// TIA Portal project "TNprojINZ" (V15.1) (continued)

       ELSIF ("OPC - z LabVIEW"."Poziom zbiornik 4" > ("OPC - do LabVIEW"."PRO poziom cieczy Z4" + 3)) THEN
           "OPC - do LabVIEW"."Zawór spustowy Z4" := 1;
           "Z4 globalne"."Czy Z4 pełny?" := 0;

       ELSIF ("OPC - z LabVIEW"."Poziom zbiornik 4" < ("OPC - do LabVIEW"."PRO poziom cieczy Z4" - 3)) THEN
           "OPC - do LabVIEW"."Zawór spustowy Z4" := 0;
           "Z4 globalne"."Czy Z4 pełny?" := 0;
       END_IF;
   //ELSE
       //"Z4 globalne"."Czy Z4 pełny?" := 0;
   END_IF;
END_FUNCTION_BLOCK

FUNCTION_BLOCK "SCL - Grzanie"   // FB9, SCL
{ S7_Optimized_Access := 'TRUE' }
VERSION : 0.1
BEGIN
   (*
   4 x - dla każdego zbiornika oddzielnie 
   if then               i Awaria = 0
       proces grzania
   else - koniec proc grz
       reset - "Z1 globalne"."Ciecz Z1 nagrzana" -> zapewniony w FB-grzałki
   *)

   // Grzałka w zbiorniku 1
   IF "Z1 globalne"."grzanie Z1 sfc" = 1 AND "Ster grzałki/zbior".HISTgrzałka1 = 1 AND "OPC - do LabVIEW".Awaria = 0
       AND "OPC - do LabVIEW"."PRO poziom cieczy Z1" >= 15 THEN
       "OPC - do LabVIEW"."Grzałka 1" := 1;
   ELSE
       "OPC - do LabVIEW"."Grzałka 1" := 0;
   END_IF;

   // Grzałka w zbiorniku 2
   IF "Z2 globalne"."grzanie Z2 sfc" = 1 AND "Ster grzałki/zbior".HISTgrzałka2 = 1 AND "OPC - do LabVIEW".Awaria = 0
       AND "OPC - do LabVIEW"."PRO poziom cieczy Z2" >= 15 THEN
       "OPC - do LabVIEW"."Grzałka 2" := 1;
   ELSE
       "OPC - do LabVIEW"."Grzałka 2" := 0;
   END_IF;

   // Grzałka w zbiorniku 3
   IF "Z3 globalne"."grzanie Z3 sfc" = 1 AND "Ster grzałki/zbior".HISTgrzałka3 = 1 AND "OPC - do LabVIEW".Awaria = 0
       AND "OPC - do LabVIEW"."PRO poziom cieczy Z3" >= 15 THEN
       "OPC - do LabVIEW"."Grzałka 3" := 1;
   ELSE
       "OPC - do LabVIEW"."Grzałka 3" := 0;
   END_IF;

   // Grzałka w zbiorniku 4
   IF "Z4 globalne"."grzanie Z4 sfc" = 1 AND "Ster grzałki/zbior".HISTgrzałka4 = 1 AND "OPC - do LabVIEW".Awaria = 0
       AND "OPC - do LabVIEW"."PRO poziom cieczy Z4" >= 15 THEN
       "OPC - do LabVIEW"."Grzałka 4" := 1;
   ELSE
       "OPC - do LabVIEW"."Grzałka 4" := 0;
   END_IF;
END_FUNCTION_BLOCK

FUNCTION_BLOCK "SCL - Awaria i zabezpieczenia par."   // FB10, SCL
{ S7_Optimized_Access := 'TRUE' }
VERSION : 0.1
BEGIN
   (*
   jak awaria = 1 to start/stop = 0
   jak awaria = 1 i poz 1-4 = 0 to wszystkie zmienne gotowości :=1
   *)
   //po awarii
   IF "Ster grzałki/zbior"."Wszystkie zbiorniki puste" = 1 AND "OPC - do LabVIEW".Awaria = 1 THEN
       "Z1 globalne"."Z1 gotowy" := 1;
       "Z2 globalne"."Z2 gotowy" := 1;
       "Z3 globalne"."Z3 gotowy" := 1;
       "Z4 globalne"."Z4 gotowy" := 1;
   END_IF;
   // reset zm proc do 0 = otwarcie zaw spust
   IF "OPC - do LabVIEW".Awaria = 1 THEN
       "HMI komunikacja"."Start/Stop" := 0;
       "OPC - do LabVIEW"."PRO poziom cieczy Z1" := 0;
       "OPC - do LabVIEW"."PRO poziom cieczy Z2" := 0;
       "OPC - do LabVIEW"."PRO poziom cieczy Z3" := 0;
       "OPC - do LabVIEW"."PRO poziom cieczy Z4" := 0;
   END_IF;
   // wyjście z stanu awaryjnego
   IF "Z1 globalne"."Awaria reset sfc Z1" = 1 AND "Z2 globalne"."Awaria reset sfc Z2" = 1 AND "Z3 globalne"."Awaria reset sfc Z3" = 1 AND
       "Z4 globalne"."Awaria reset sfc Z4" = 1 THEN
       "OPC - do LabVIEW".Awaria := 0;
       "OPC - do LabVIEW"."Zawór spustowy Z1" := 0;
       "OPC - do LabVIEW"."Zawór spustowy Z2" := 0;
       "OPC - do LabVIEW"."Zawór spustowy Z3" := 0;
       "OPC - do LabVIEW"."Zawór spustowy Z4" := 0;
   END_IF;

   IF "Z1 globalne"."Awaria reset sfc Z1" = 1 THEN
       "OPC - do LabVIEW"."PRO poziom cieczy Z1" := 0;
   END_IF;

   IF "Z2 globalne"."Awaria reset sfc Z2" = 1 THEN
       "OPC - do LabVIEW"."PRO poziom cieczy Z2" := 0;
   END_IF;

   IF "Z3 globalne"."Awaria reset sfc Z3" = 1 THEN
       "OPC - do LabVIEW"."PRO poziom cieczy Z3" := 0;
   END_IF;

   //Zabezpieczenie parametrów procesu wybranych w HMI
   //Z1
   IF "HMI komunikacja"."HMI poziom cieczy Z1" < 15 THEN
       "HMI komunikacja"."HMI poziom cieczy Z1" := 0;
       "HMI komunikacja"."HMI czas utrz T  Z1" := 0;
       "HMI komunikacja"."HMI Temp max Z1" := 20;
   END_IF;

   IF "HMI komunikacja"."HMI Temp max Z1" < 40 THEN
       "HMI komunikacja"."HMI Temp max Z1" := 20;
   END_IF;

   IF "HMI komunikacja"."HMI czas utrz T  Z1" < 5 THEN
       "HMI komunikacja"."HMI czas utrz T  Z1" := 0;
   END_IF;

   //Z2
   IF "HMI komunikacja"."HMI poziom cieczy Z2" < 15 THEN
       "HMI komunikacja"."HMI poziom cieczy Z2" := 0;
       "HMI komunikacja"."HMI czas utrz T  Z2" := 0;
       "HMI komunikacja"."HMI Temp max Z2" := 20;
   END_IF;

   IF "HMI komunikacja"."HMI Temp max Z2" < 40 THEN
       "HMI komunikacja"."HMI Temp max Z2" := 20;
   END_IF;

   IF "HMI komunikacja"."HMI czas utrz T  Z2" < 5 THEN
       "HMI komunikacja"."HMI czas utrz T  Z2" := 0;
   END_IF;

   //Z3
   IF "HMI komunikacja"."HMI poziom cieczy Z3" < 15 THEN
       "HMI komunikacja"."HMI poziom cieczy Z3" := 0;
       "HMI komunikacja"."HMI czas utrz T  Z3" := 0;
       "HMI komunikacja"."HMI Temp max Z3" := 20;
   END_IF;

   IF "HMI komunikacja"."HMI Temp max Z3" < 40 THEN
       "HMI komunikacja"."HMI Temp max Z3" := 20;
   END_IF;

   IF "HMI komunikacja"."HMI czas utrz T  Z3" < 5 THEN
       "HMI komunikacja"."HMI czas utrz T  Z3" := 0;
   END_IF;

   //Z4
   IF "HMI komunikacja"."HMI Temp max Z4" < 40 THEN
       "HMI komunikacja"."HMI Temp max Z4" := 20;
   END_IF;

   IF "HMI komunikacja"."HMI czas utrz T  Z4" < 5 THEN
       "HMI komunikacja"."HMI czas utrz T  Z4" := 0;
   END_IF;
END_FUNCTION_BLOCK

FUNCTION_BLOCK "FB - pompy"   // FB11, FBD
{ S7_Optimized_Access := 'TRUE' }
VERSION : 0.1
BEGIN

REGION Network 1: Pompy P1-P2 przegrzane
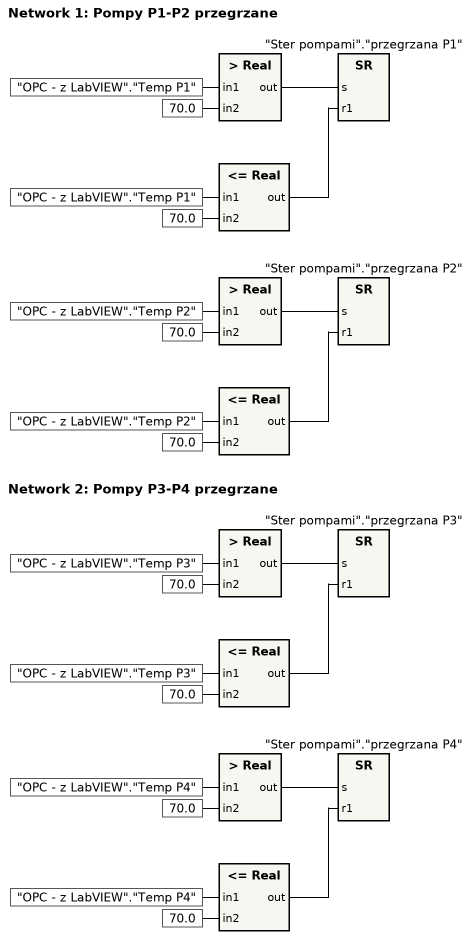
   IF "OPC - z LabVIEW"."Temp P1" > 70.0 THEN
       "Ster pompami"."przegrzana P1" := TRUE;   // SR flip-flop
   END_IF;
   IF "OPC - z LabVIEW"."Temp P1" <= 70.0 THEN "Ster pompami"."przegrzana P1" := FALSE; END_IF;
   IF "OPC - z LabVIEW"."Temp P2" > 70.0 THEN
       "Ster pompami"."przegrzana P2" := TRUE;   // SR flip-flop
   END_IF;
   IF "OPC - z LabVIEW"."Temp P2" <= 70.0 THEN "Ster pompami"."przegrzana P2" := FALSE; END_IF;
END_REGION

REGION Network 2: Pompy P3-P4 przegrzane
   IF "OPC - z LabVIEW"."Temp P3" > 70.0 THEN
       "Ster pompami"."przegrzana P3" := TRUE;   // SR flip-flop
   END_IF;
   IF "OPC - z LabVIEW"."Temp P3" <= 70.0 THEN "Ster pompami"."przegrzana P3" := FALSE; END_IF;
   IF "OPC - z LabVIEW"."Temp P4" > 70.0 THEN
       "Ster pompami"."przegrzana P4" := TRUE;   // SR flip-flop
   END_IF;
   IF "OPC - z LabVIEW"."Temp P4" <= 70.0 THEN "Ster pompami"."przegrzana P4" := FALSE; END_IF;
END_REGION

REGION Network 3: Pompy P5-P6 przegrzane
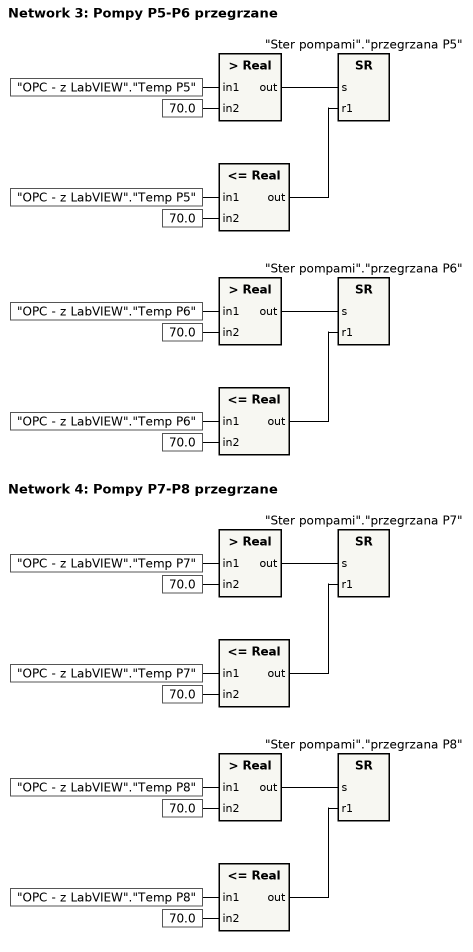
   IF "OPC - z LabVIEW"."Temp P5" > 70.0 THEN
       "Ster pompami"."przegrzana P5" := TRUE;   // SR flip-flop
   END_IF;
   IF "OPC - z LabVIEW"."Temp P5" <= 70.0 THEN "Ster pompami"."przegrzana P5" := FALSE; END_IF;
   IF "OPC - z LabVIEW"."Temp P6" > 70.0 THEN
       "Ster pompami"."przegrzana P6" := TRUE;   // SR flip-flop
   END_IF;
   IF "OPC - z LabVIEW"."Temp P6" <= 70.0 THEN "Ster pompami"."przegrzana P6" := FALSE; END_IF;
END_REGION

REGION Network 4: Pompy P7-P8 przegrzane
   IF "OPC - z LabVIEW"."Temp P7" > 70.0 THEN
       "Ster pompami"."przegrzana P7" := TRUE;   // SR flip-flop
   END_IF;
   IF "OPC - z LabVIEW"."Temp P7" <= 70.0 THEN "Ster pompami"."przegrzana P7" := FALSE; END_IF;
   IF "OPC - z LabVIEW"."Temp P8" > 70.0 THEN
       "Ster pompami"."przegrzana P8" := TRUE;   // SR flip-flop
   END_IF;
   IF "OPC - z LabVIEW"."Temp P8" <= 70.0 THEN "Ster pompami"."przegrzana P8" := FALSE; END_IF;
END_REGION
END_FUNCTION_BLOCK

ORGANIZATION_BLOCK "Main"   // OB1, LAD, ProgramCycle
TITLE = "Main Program Sweep (Cycle)"
{ S7_Optimized_Access := 'TRUE' }
VERSION : 0.1
   VAR_INPUT
      Initial_Call : Bool;   // Initial call of this OB
      Remanence : Bool;   // =True, if remanent data are available
   END_VAR
BEGIN

REGION Network 1: SFC - Zbiornik 1
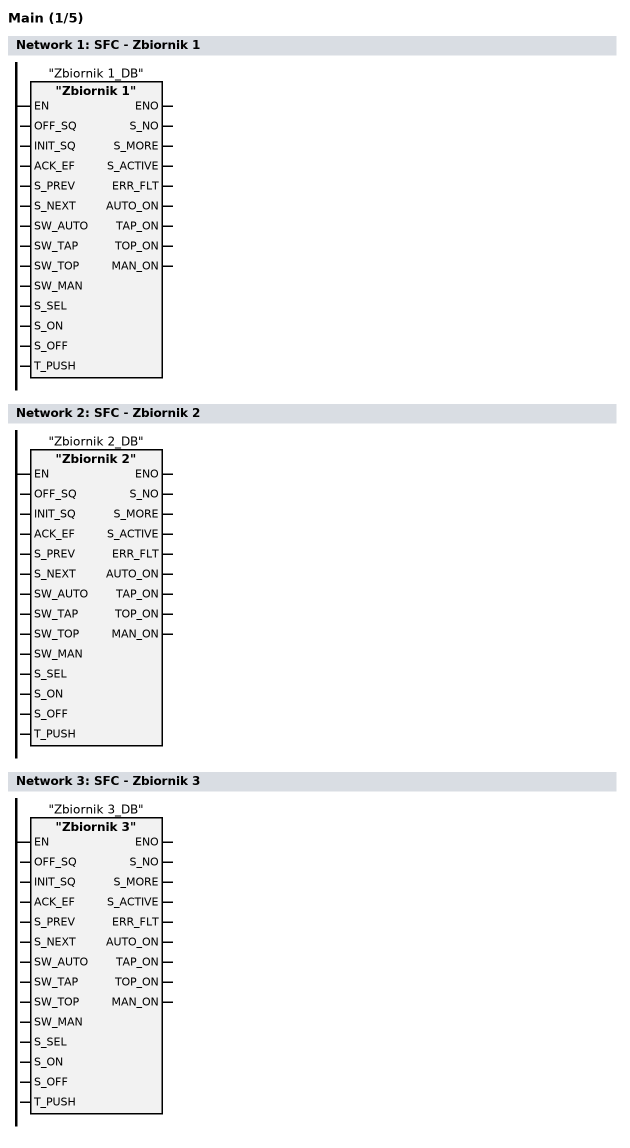
   RUNG wire#powerrail
      "Zbiornik 1_DB"(OFF_SQ :=, INIT_SQ :=, ACK_EF :=, S_PREV :=, S_NEXT :=, SW_AUTO :=, SW_TAP :=, SW_TOP :=, SW_MAN :=, S_SEL :=, S_ON :=, S_OFF :=, T_PUSH :=, S_NO =>, S_MORE =>, S_ACTIVE =>, ERR_FLT =>, AUTO_ON =>, TAP_ON =>, TOP_ON =>, MAN_ON =>)
   END_RUNG
   // the same network as SCL:
   "Zbiornik 1_DB"();   // "Zbiornik 1"
END_REGION

REGION Network 2: SFC - Zbiornik 2
   RUNG wire#powerrail
      "Zbiornik 2_DB"(OFF_SQ :=, INIT_SQ :=, ACK_EF :=, S_PREV :=, S_NEXT :=, SW_AUTO :=, SW_TAP :=, SW_TOP :=, SW_MAN :=, S_SEL :=, S_ON :=, S_OFF :=, T_PUSH :=, S_NO =>, S_MORE =>, S_ACTIVE =>, ERR_FLT =>, AUTO_ON =>, TAP_ON =>, TOP_ON =>, MAN_ON =>)
   END_RUNG
   // the same network as SCL:
   "Zbiornik 2_DB"();   // "Zbiornik 2"
END_REGION

REGION Network 3: SFC - Zbiornik 3
   RUNG wire#powerrail
      "Zbiornik 3_DB"(OFF_SQ :=, INIT_SQ :=, ACK_EF :=, S_PREV :=, S_NEXT :=, SW_AUTO :=, SW_TAP :=, SW_TOP :=, SW_MAN :=, S_SEL :=, S_ON :=, S_OFF :=, T_PUSH :=, S_NO =>, S_MORE =>, S_ACTIVE =>, ERR_FLT =>, AUTO_ON =>, TAP_ON =>, TOP_ON =>, MAN_ON =>)
   END_RUNG
   // the same network as SCL:
   "Zbiornik 3_DB"();   // "Zbiornik 3"
END_REGION

REGION Network 4: SFC - Zbiornik 4
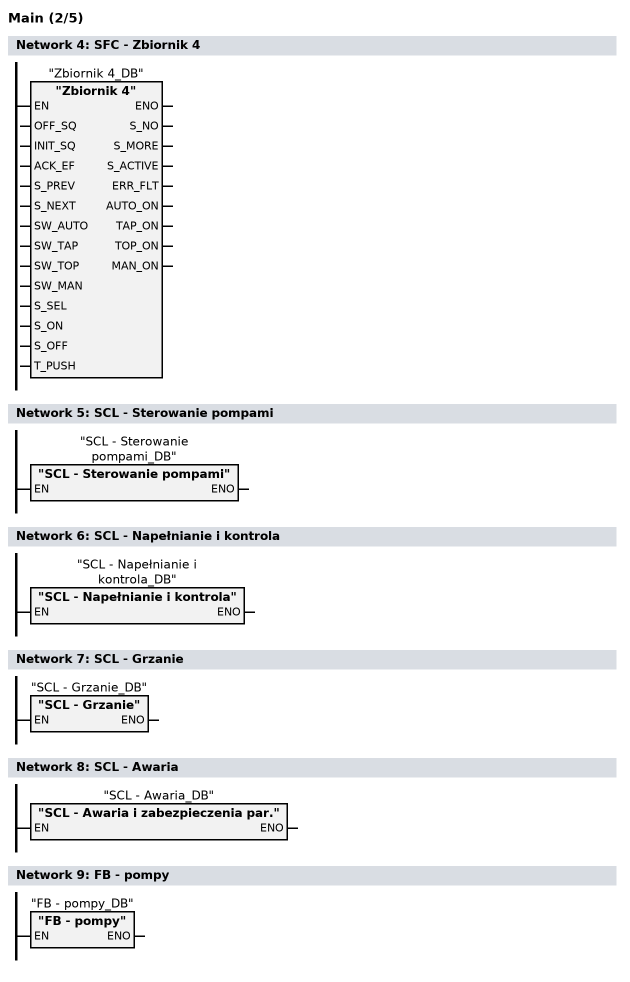
   RUNG wire#powerrail
      "Zbiornik 4_DB"(OFF_SQ :=, INIT_SQ :=, ACK_EF :=, S_PREV :=, S_NEXT :=, SW_AUTO :=, SW_TAP :=, SW_TOP :=, SW_MAN :=, S_SEL :=, S_ON :=, S_OFF :=, T_PUSH :=, S_NO =>, S_MORE =>, S_ACTIVE =>, ERR_FLT =>, AUTO_ON =>, TAP_ON =>, TOP_ON =>, MAN_ON =>)
   END_RUNG
   // the same network as SCL:
   "Zbiornik 4_DB"();   // "Zbiornik 4"
END_REGION

REGION Network 5: SCL - Sterowanie pompami
   RUNG wire#powerrail
      "SCL - Sterowanie pompami_DB"()
   END_RUNG
   // the same network as SCL:
   "SCL - Sterowanie pompami_DB"();   // "SCL - Sterowanie pompami"
END_REGION

REGION Network 6: SCL - Napełnianie i kontrola
   RUNG wire#powerrail
      "SCL - Napełnianie i kontrola_DB"()
   END_RUNG
   // the same network as SCL:
   "SCL - Napełnianie i kontrola_DB"();   // "SCL - Napełnianie i kontrola"
END_REGION

REGION Network 7: SCL - Grzanie
   RUNG wire#powerrail
      "SCL - Grzanie_DB"()
   END_RUNG
   // the same network as SCL:
   "SCL - Grzanie_DB"();   // "SCL - Grzanie"
END_REGION

REGION Network 8: SCL - Awaria
   RUNG wire#powerrail
      "SCL - Awaria_DB"()
   END_RUNG
   // the same network as SCL:
   "SCL - Awaria_DB"();   // "SCL - Awaria i zabezpieczenia par."
END_REGION

REGION Network 9: FB - pompy
   RUNG wire#powerrail
      "FB - pompy_DB"()
   END_RUNG
   // the same network as SCL:
   "FB - pompy_DB"();   // "FB - pompy"
END_REGION

REGION Network 10: FB - grzałki
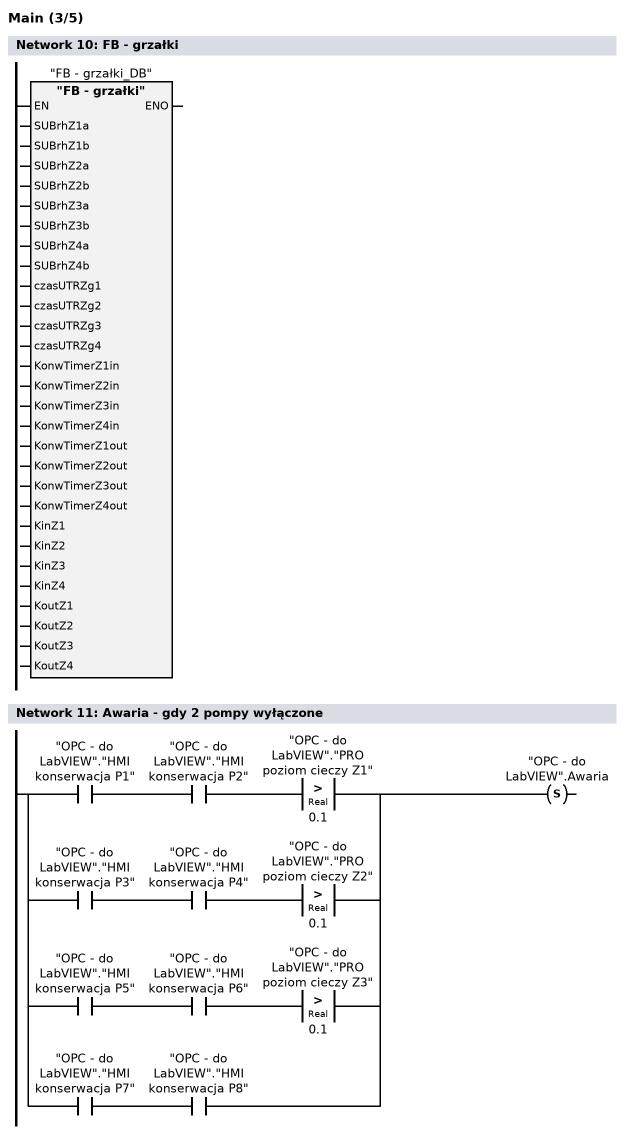
   RUNG wire#powerrail
      "FB - grzałki_DB"(SUBrhZ1a :=, SUBrhZ1b :=, SUBrhZ2a :=, SUBrhZ2b :=, SUBrhZ3a :=, SUBrhZ3b :=, SUBrhZ4a :=, SUBrhZ4b :=, czasUTRZg1 :=, czasUTRZg2 :=, czasUTRZg3 :=, czasUTRZg4 :=, KonwTimerZ1in :=, KonwTimerZ2in :=, KonwTimerZ3in :=, KonwTimerZ4in :=, KonwTimerZ1out :=, KonwTimerZ2out :=, KonwTimerZ3out :=, KonwTimerZ4out :=, KinZ1 :=, KinZ2 :=, KinZ3 :=, KinZ4 :=, KoutZ1 :=, KoutZ2 :=, KoutZ3 :=, KoutZ4 :=)
   END_RUNG
   // the same network as SCL:
   "FB - grzałki_DB"();   // "FB - grzałki"
END_REGION

REGION Network 11: Awaria - gdy 2 pompy wyłączone
   RUNG wire#powerrail
      Contact( "OPC - do LabVIEW"."HMI konserwacja P1" )
      Contact( "OPC - do LabVIEW"."HMI konserwacja P2" )
      { S7_Templates := "SrcType := Real" } GT_Contact(in1 := "OPC - do LabVIEW"."PRO poziom cieczy Z1", in2 := 0.1)
      wire#w1
      S_Coil( "OPC - do LabVIEW".Awaria )
   END_RUNG
   RUNG wire#powerrail
      Contact( "OPC - do LabVIEW"."HMI konserwacja P3" )
      Contact( "OPC - do LabVIEW"."HMI konserwacja P4" )
      { S7_Templates := "SrcType := Real" } GT_Contact(in1 := "OPC - do LabVIEW"."PRO poziom cieczy Z2", in2 := 0.1)
   END_RUNG wire#w1
   RUNG wire#powerrail
      Contact( "OPC - do LabVIEW"."HMI konserwacja P5" )
      Contact( "OPC - do LabVIEW"."HMI konserwacja P6" )
      { S7_Templates := "SrcType := Real" } GT_Contact(in1 := "OPC - do LabVIEW"."PRO poziom cieczy Z3", in2 := 0.1)
   END_RUNG wire#w1
   RUNG wire#powerrail
      Contact( "OPC - do LabVIEW"."HMI konserwacja P7" )
      Contact( "OPC - do LabVIEW"."HMI konserwacja P8" )
   END_RUNG wire#w1
   // the same network as SCL:
   IF ("OPC - do LabVIEW"."HMI konserwacja P1" AND "OPC - do LabVIEW"."HMI konserwacja P2" AND ("OPC - do LabVIEW"."PRO poziom cieczy Z1" > 0.1)) OR ("OPC - do LabVIEW"."HMI konserwacja P3" AND "OPC - do LabVIEW"."HMI konserwacja P4" AND ("OPC - do LabVIEW"."PRO poziom cieczy Z2" > 0.1)) OR ("OPC - do LabVIEW"."HMI konserwacja P5" AND "OPC - do LabVIEW"."HMI konserwacja P6" AND ("OPC - do LabVIEW"."PRO poziom cieczy Z3" > 0.1)) OR ("OPC - do LabVIEW"."HMI konserwacja P7" AND "OPC - do LabVIEW"."HMI konserwacja P8") THEN
       "OPC - do LabVIEW".Awaria := TRUE;
   END_IF;
END_REGION

REGION Network 12: Załączenie zaworów spustowych podczas Awarii
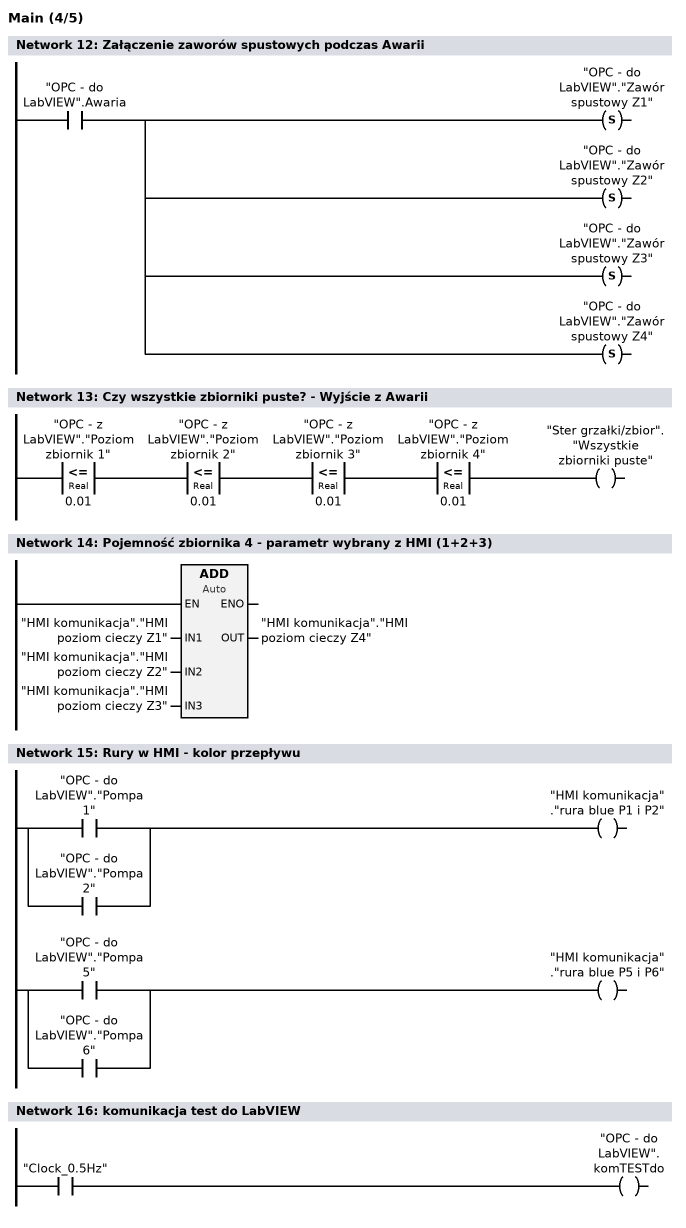
   RUNG wire#powerrail
      Contact( "OPC - do LabVIEW".Awaria )
      wire#w1
      S_Coil( "OPC - do LabVIEW"."Zawór spustowy Z1" )
   END_RUNG
   RUNG wire#w1
      S_Coil( "OPC - do LabVIEW"."Zawór spustowy Z2" )
   END_RUNG
   RUNG wire#w1
      S_Coil( "OPC - do LabVIEW"."Zawór spustowy Z3" )
   END_RUNG
   RUNG wire#w1
      S_Coil( "OPC - do LabVIEW"."Zawór spustowy Z4" )
   END_RUNG
   // the same network as SCL:
   IF "OPC - do LabVIEW".Awaria THEN
       "OPC - do LabVIEW"."Zawór spustowy Z1" := TRUE;
       "OPC - do LabVIEW"."Zawór spustowy Z2" := TRUE;
       "OPC - do LabVIEW"."Zawór spustowy Z3" := TRUE;
       "OPC - do LabVIEW"."Zawór spustowy Z4" := TRUE;
   END_IF;
END_REGION

REGION Network 13: Czy wszystkie zbiorniki puste? - Wyjście z Awarii
   RUNG wire#powerrail
      { S7_Templates := "SrcType := Real" } LE_Contact(in1 := "OPC - z LabVIEW"."Poziom zbiornik 1", in2 := 0.01)
      { S7_Templates := "SrcType := Real" } LE_Contact(in1 := "OPC - z LabVIEW"."Poziom zbiornik 2", in2 := 0.01)
      { S7_Templates := "SrcType := Real" } LE_Contact(in1 := "OPC - z LabVIEW"."Poziom zbiornik 3", in2 := 0.01)
      { S7_Templates := "SrcType := Real" } LE_Contact(in1 := "OPC - z LabVIEW"."Poziom zbiornik 4", in2 := 0.01)
      Coil( "Ster grzałki/zbior"."Wszystkie zbiorniki puste" )
   END_RUNG
   // the same network as SCL:
   "Ster grzałki/zbior"."Wszystkie zbiorniki puste" := ("OPC - z LabVIEW"."Poziom zbiornik 1" <= 0.01) AND ("OPC - z LabVIEW"."Poziom zbiornik 2" <= 0.01) AND ("OPC - z LabVIEW"."Poziom zbiornik 3" <= 0.01) AND ("OPC - z LabVIEW"."Poziom zbiornik 4" <= 0.01);
END_REGION

REGION Network 14: Pojemność zbiornika 4 - parametr wybrany z HMI (1+2+3)
   RUNG wire#powerrail
      Add(in1 := "HMI komunikacja"."HMI poziom cieczy Z1", in2 := "HMI komunikacja"."HMI poziom cieczy Z2", in3 := "HMI komunikacja"."HMI poziom cieczy Z3", out => "HMI komunikacja"."HMI poziom cieczy Z4")
   END_RUNG
   // the same network as SCL:
   "HMI komunikacja"."HMI poziom cieczy Z4" := "HMI komunikacja"."HMI poziom cieczy Z1" + "HMI komunikacja"."HMI poziom cieczy Z2" + "HMI komunikacja"."HMI poziom cieczy Z3";
END_REGION

REGION Network 15: Rury w HMI - kolor przepływu
   RUNG wire#powerrail
      Contact( "OPC - do LabVIEW"."Pompa 1" )
      wire#w1
      Coil( "HMI komunikacja"."rura blue P1 i P2" )
   END_RUNG
   RUNG wire#powerrail
      Contact( "OPC - do LabVIEW"."Pompa 2" )
   END_RUNG wire#w1
   RUNG wire#powerrail
      Contact( "OPC - do LabVIEW"."Pompa 5" )
      wire#w2
      Coil( "HMI komunikacja"."rura blue P5 i P6" )
   END_RUNG
   RUNG wire#powerrail
      Contact( "OPC - do LabVIEW"."Pompa 6" )
   END_RUNG wire#w2
   // the same network as SCL:
   "HMI komunikacja"."rura blue P1 i P2" := "OPC - do LabVIEW"."Pompa 1" OR "OPC - do LabVIEW"."Pompa 2";
   "HMI komunikacja"."rura blue P5 i P6" := "OPC - do LabVIEW"."Pompa 5" OR "OPC - do LabVIEW"."Pompa 6";
END_REGION

REGION Network 16: komunikacja test do LabVIEW
   RUNG wire#powerrail
      Contact( "Clock_0.5Hz" )
      Coil( "OPC - do LabVIEW".komTESTdo )
   END_RUNG
   // the same network as SCL:
   "OPC - do LabVIEW".komTESTdo := "Clock_0.5Hz";
END_REGION

REGION Network 17: komunikacja test z LabVIEW
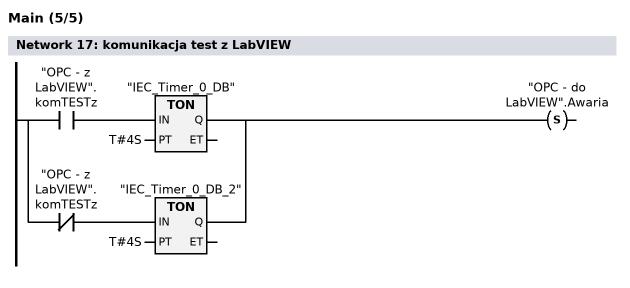
   "IEC_Timer_0_DB".TON(IN := "OPC - z LabVIEW".komTESTz, PT := T#4S);
   "IEC_Timer_0_DB_2".TON(IN := NOT "OPC - z LabVIEW".komTESTz, PT := T#4S);
   IF "IEC_Timer_0_DB".Q OR "IEC_Timer_0_DB_2".Q THEN "OPC - do LabVIEW".Awaria := TRUE; END_IF;
END_REGION
END_ORGANIZATION_BLOCK

(* ===== HMI "HMI_RT_1" =====
system functions are stored by id; their names below are inferred from use
connection "HMI_Connection_2": ETHERNET, S7_1500_OMS

HMI tags "Default tag table"
   "Clock_1Hz" : Bool = PLC Clock_1Hz AT %M0.5, 100 ms
   "Clock_0.5Hz" : Bool = PLC "Clock_0.5Hz" AT %M0.7, 100 ms
   "HMI komunikacja_Start/Stop" : Bool = PLC "HMI komunikacja".Start/Stop AT %DB2.DBX0.0, 100 ms
   "OPC - do LabVIEW_Awaria" : Bool = PLC "OPC - do LabVIEW".Awaria AT %DB4.DBX48.0, 100 ms
   "OPC - do LabVIEW_Pompa 1" : Bool = PLC "OPC - do LabVIEW"."Pompa 1" AT %DB4.DBX48.1, 100 ms
   "OPC - z LabVIEW_Temp P1" : Real = PLC "OPC - z LabVIEW"."Temp P1" AT %DB3.DBD0, 100 ms
   "OPC - do LabVIEW_HMI konserwacja P1" : Bool = PLC "OPC - do LabVIEW"."HMI konserwacja P1" AT %DB4.DBX50.0, 100 ms
   "OPC - do LabVIEW_HMI konserwacja P2" : Bool = PLC "OPC - do LabVIEW"."HMI konserwacja P2" AT %DB4.DBX50.1, 100 ms
   "OPC - do LabVIEW_HMI konserwacja P3" : Bool = PLC "OPC - do LabVIEW"."HMI konserwacja P3" AT %DB4.DBX50.2, 100 ms
   "OPC - do LabVIEW_HMI konserwacja P4" : Bool = PLC "OPC - do LabVIEW"."HMI konserwacja P4" AT %DB4.DBX50.3, 100 ms
   "OPC - do LabVIEW_HMI konserwacja P5" : Bool = PLC "OPC - do LabVIEW"."HMI konserwacja P5" AT %DB4.DBX50.4, 100 ms
   "OPC - do LabVIEW_HMI konserwacja P6" : Bool = PLC "OPC - do LabVIEW"."HMI konserwacja P6" AT %DB4.DBX50.5, 100 ms
   "OPC - do LabVIEW_HMI konserwacja P7" : Bool = PLC "OPC - do LabVIEW"."HMI konserwacja P7" AT %DB4.DBX50.6, 100 ms
   "OPC - do LabVIEW_HMI konserwacja P8" : Bool = PLC "OPC - do LabVIEW"."HMI konserwacja P8" AT %DB4.DBX50.7, 100 ms
   "OPC - do LabVIEW_Zawór wlotowy 1" : Bool = PLC "OPC - do LabVIEW"."Zawór wlotowy 1" AT %DB4.DBX49.1, 100 ms
   "OPC - do LabVIEW_Zawór wlotowy 2" : Bool = PLC "OPC - do LabVIEW"."Zawór wlotowy 2" AT %DB4.DBX49.2, 100 ms
   "OPC - do LabVIEW_Zawór wlotowy 3" : Bool = PLC "OPC - do LabVIEW"."Zawór wlotowy 3" AT %DB4.DBX49.3, 100 ms
   "OPC - z LabVIEW_Temp cieczy w zb1" : Real = PLC "OPC - z LabVIEW"."Temp cieczy w zb1" AT %DB3.DBD32, 100 ms
   "OPC - z LabVIEW_Temp cieczy w zb2" : Real = PLC "OPC - z LabVIEW"."Temp cieczy w zb2" AT %DB3.DBD36, 100 ms
   "OPC - z LabVIEW_Temp cieczy w zb3" : Real = PLC "OPC - z LabVIEW"."Temp cieczy w zb3" AT %DB3.DBD40, 100 ms
   "OPC - z LabVIEW_Temp cieczy w zb4" : Real = PLC "OPC - z LabVIEW"."Temp cieczy w zb4" AT %DB3.DBD44, 100 ms
   "HMI komunikacja_Czas utrz T w Z1 (timer)" : Real = PLC "HMI komunikacja"."Czas utrz T w Z1 (timer)", 100 ms
   "HMI komunikacja_Czas utrz T w Z2 (timer)" : Real = PLC "HMI komunikacja"."Czas utrz T w Z2 (timer)", 100 ms
   "HMI komunikacja_Czas utrz T w Z3 (timer)" : Real = PLC "HMI komunikacja"."Czas utrz T w Z3 (timer)", 100 ms
   "HMI komunikacja_Czas utrz T w Z4 (timer)" : Real = PLC "HMI komunikacja"."Czas utrz T w Z4 (timer)", 100 ms
   "OPC - do LabVIEW_Grzałka 1" : Bool = PLC "OPC - do LabVIEW"."Grzałka 1" AT %DB4.DBX49.4, 100 ms
   "OPC - do LabVIEW_Grzałka 2" : Bool = PLC "OPC - do LabVIEW"."Grzałka 2" AT %DB4.DBX49.5, 100 ms
   "OPC - do LabVIEW_Grzałka 3" : Bool = PLC "OPC - do LabVIEW"."Grzałka 3" AT %DB4.DBX49.6, 100 ms
   "OPC - do LabVIEW_Grzałka 4" : Bool = PLC "OPC - do LabVIEW"."Grzałka 4" AT %DB4.DBX49.7, 100 ms
   "OPC - do LabVIEW_Pompa 2" : Bool = PLC "OPC - do LabVIEW"."Pompa 2" AT %DB4.DBX48.2, 100 ms
   "OPC - do LabVIEW_Pompa 3" : Bool = PLC "OPC - do LabVIEW"."Pompa 3" AT %DB4.DBX48.3, 100 ms
   "OPC - do LabVIEW_Pompa 4" : Bool = PLC "OPC - do LabVIEW"."Pompa 4" AT %DB4.DBX48.4, 100 ms
   "OPC - do LabVIEW_Pompa 5" : Bool = PLC "OPC - do LabVIEW"."Pompa 5" AT %DB4.DBX48.5, 100 ms
   "OPC - do LabVIEW_Pompa 6" : Bool = PLC "OPC - do LabVIEW"."Pompa 6" AT %DB4.DBX48.6, 100 ms
   "OPC - do LabVIEW_Pompa 7" : Bool = PLC "OPC - do LabVIEW"."Pompa 7" AT %DB4.DBX48.7, 100 ms
   "OPC - do LabVIEW_Pompa 8" : Bool = PLC "OPC - do LabVIEW"."Pompa 8" AT %DB4.DBX49.0, 100 ms
   "OPC - z LabVIEW_Temp P2" : Real = PLC "OPC - z LabVIEW"."Temp P2" AT %DB3.DBD4, 100 ms
   "OPC - z LabVIEW_Temp P3" : Real = PLC "OPC - z LabVIEW"."Temp P3" AT %DB3.DBD8, 100 ms
   "OPC - z LabVIEW_Temp P4" : Real = PLC "OPC - z LabVIEW"."Temp P4" AT %DB3.DBD12, 100 ms
   "OPC - z LabVIEW_Temp P5" : Real = PLC "OPC - z LabVIEW"."Temp P5" AT %DB3.DBD16, 100 ms
   "OPC - z LabVIEW_Temp P6" : Real = PLC "OPC - z LabVIEW"."Temp P6" AT %DB3.DBD20, 100 ms
   "OPC - z LabVIEW_Temp P7" : Real = PLC "OPC - z LabVIEW"."Temp P7" AT %DB3.DBD24, 100 ms
   "OPC - z LabVIEW_Temp P8" : Real = PLC "OPC - z LabVIEW"."Temp P8" AT %DB3.DBD28, 100 ms
   "HMI komunikacja_rura blue P1 i P2" : Bool = PLC "HMI komunikacja"."rura blue P1 i P2", 100 ms
   "HMI komunikacja_rura blue P5 i P6" : Bool = PLC "HMI komunikacja"."rura blue P5 i P6", 100 ms
   "HMI komunikacja_HMI poziom cieczy Z1" : Real = PLC "HMI komunikacja"."HMI poziom cieczy Z1", 100 ms
   "HMI komunikacja_HMI poziom cieczy Z2" : Real = PLC "HMI komunikacja"."HMI poziom cieczy Z2", 100 ms
   "HMI komunikacja_HMI poziom cieczy Z3" : Real = PLC "HMI komunikacja"."HMI poziom cieczy Z3", 100 ms
   "HMI komunikacja_HMI poziom cieczy Z4" : Real = PLC "HMI komunikacja"."HMI poziom cieczy Z4", 100 ms
   "HMI komunikacja_HMI Temp max Z1" : Real = PLC "HMI komunikacja"."HMI Temp max Z1", 100 ms
   "HMI komunikacja_HMI Temp max Z2" : Real = PLC "HMI komunikacja"."HMI Temp max Z2", 100 ms
   "HMI komunikacja_HMI Temp max Z3" : Real = PLC "HMI komunikacja"."HMI Temp max Z3", 100 ms
   "HMI komunikacja_HMI czas utrz T  Z1" : Real = PLC "HMI komunikacja"."HMI czas utrz T  Z1", 100 ms
   "HMI komunikacja_HMI czas utrz T  Z2" : Real = PLC "HMI komunikacja"."HMI czas utrz T  Z2", 100 ms
   "HMI komunikacja_HMI czas utrz T  Z3" : Real = PLC "HMI komunikacja"."HMI czas utrz T  Z3", 100 ms
   "HMI komunikacja_HMI Temp max Z4" : Real = PLC "HMI komunikacja"."HMI Temp max Z4", 100 ms
   "HMI komunikacja_HMI czas utrz T  Z4" : Real = PLC "HMI komunikacja"."HMI czas utrz T  Z4", 100 ms
   "OPC - do LabVIEW_Zawór spustowy Z4" : Bool = PLC "OPC - do LabVIEW"."Zawór spustowy Z4" AT %DB4.DBX51.3, 100 ms
   "OPC - do LabVIEW_Zawór spustowy Z1" : Bool = PLC "OPC - do LabVIEW"."Zawór spustowy Z1" AT %DB4.DBX51.0, 100 ms
   "OPC - do LabVIEW_Zawór spustowy Z2" : Bool = PLC "OPC - do LabVIEW"."Zawór spustowy Z2" AT %DB4.DBX51.1, 100 ms
   "OPC - do LabVIEW_Zawór spustowy Z3" : Bool = PLC "OPC - do LabVIEW"."Zawór spustowy Z3" AT %DB4.DBX51.2, 100 ms
   "OPC - z LabVIEW_Poziom zbiornik 1" : Real = PLC "OPC - z LabVIEW"."Poziom zbiornik 1" AT %DB3.DBD48, 100 ms
   "OPC - z LabVIEW_Poziom zbiornik 2" : Real = PLC "OPC - z LabVIEW"."Poziom zbiornik 2" AT %DB3.DBD52, 100 ms
   "OPC - z LabVIEW_Poziom zbiornik 3" : Real = PLC "OPC - z LabVIEW"."Poziom zbiornik 3" AT %DB3.DBD56, 100 ms
   "OPC - z LabVIEW_Poziom zbiornik 4" : Real = PLC "OPC - z LabVIEW"."Poziom zbiornik 4" AT %DB3.DBD60, 100 ms
   "HMI komunikacja_Blokada zmiany par. PRO" : Bool = PLC "HMI komunikacja"."Blokada zmiany par. PRO", 1 s

screen "Wizualizacja i start" 800x434
   SymbolLibrary "Symbol library_4" at 337,36 size 132x115
   TextField "Text field_1" at 0,0 size 149x18; Text 'Wizualizacja procesu'
   SymbolLibrary "Symbol library_1" at 384,0 size 31x37
      Appearance <- "OPC - do LabVIEW_Zawór wlotowy 2"
   Bar "Bar_1" at 338,37 size 38x113; MinimumValue 0; MaximumValue 100
      ProcessValue <- "OPC - z LabVIEW_Poziom zbiornik 2"
   SymbolLibrary "Symbol library_2" at 361,372 size 28x45
      Appearance <- "OPC - do LabVIEW_Pompa 7"
   SymbolLibrary "Symbol library_3" at 363,416 size 16x18
      Appearance <- "OPC - do LabVIEW_Pompa 7"
   SymbolLibrary "Symbol library_7" at 227,258 size 345x115
   SymbolLibrary "Symbol library_8" at 175,0 size 31x37
      Appearance <- "OPC - do LabVIEW_Zawór wlotowy 1"
   SymbolLibrary "Symbol library_9" at 599,0 size 31x37
      Appearance <- "OPC - do LabVIEW_Zawór wlotowy 3"
   SymbolLibrary "Symbol library_10" at 385,130 size 62x20
      Appearance <- "OPC - do LabVIEW_Grzałka 2"
   IOField "I/O field_1" at 379,40 size 48x31; FormatPattern 999
      ProcessValue <- "HMI komunikacja_Czas utrz T w Z2 (timer)"
   IOField "I/O field_2" at 377,98 size 70x31; FormatPattern 999.9
      ProcessValue <- "OPC - z LabVIEW_Temp cieczy w zb2"
   TextField "Text field_2" at 435,54 size 33x18; Text 'sek.'
   TextField "Text field_3" at 442,107 size 25x23; Text '℃'
   SymbolLibrary "Symbol library_6" at 127,36 size 132x115
   Bar "Bar_2" at 128,37 size 38x113; MinimumValue 0; MaximumValue 100
      ProcessValue <- "OPC - z LabVIEW_Poziom zbiornik 1"
   SymbolLibrary "Symbol library_11" at 175,130 size 62x20
      Appearance <- "OPC - do LabVIEW_Grzałka 1"
   IOField "I/O field_3" at 169,40 size 48x31; FormatPattern 999
      ProcessValue <- "HMI komunikacja_Czas utrz T w Z1 (timer)"
   IOField "I/O field_4" at 167,98 size 70x31; FormatPattern 999.9
      ProcessValue <- "OPC - z LabVIEW_Temp cieczy w zb1"
   TextField "Text field_4" at 225,54 size 33x18; Text 'sek.'
   TextField "Text field_5" at 233,107 size 25x23; Text '℃'
   SymbolLibrary "Symbol library_12" at 548,36 size 132x115
   Bar "Bar_3" at 549,37 size 38x113; MinimumValue 0; MaximumValue 100
      ProcessValue <- "OPC - z LabVIEW_Poziom zbiornik 3"
   SymbolLibrary "Symbol library_13" at 596,130 size 62x20
      Appearance <- "OPC - do LabVIEW_Grzałka 3"
   IOField "I/O field_5" at 590,40 size 48x31; FormatPattern 999
      ProcessValue <- "HMI komunikacja_Czas utrz T w Z3 (timer)"
   IOField "I/O field_6" at 588,98 size 70x31; FormatPattern 999.9
      ProcessValue <- "OPC - z LabVIEW_Temp cieczy w zb3"
   TextField "Text field_6" at 646,54 size 33x18; Text 'sek.'
   TextField "Text field_7" at 654,107 size 25x23; Text '℃'
   SymbolLibrary "Symbol library_14" at 151,165 size 28x45
      Appearance <- "OPC - do LabVIEW_Pompa 1"
   SymbolLibrary "Symbol library_15" at 152,151 size 16x15
      Appearance <- "OPC - do LabVIEW_Pompa 1"
   SymbolLibrary "Symbol library_5" at 197,165 size 28x45
      Appearance <- "OPC - do LabVIEW_Pompa 2"
   SymbolLibrary "Symbol library_16" at 198,151 size 16x15
      Appearance <- "OPC - do LabVIEW_Pompa 2"
   SymbolLibrary "Symbol library_17" at 360,165 size 28x45
      Appearance <- "OPC - do LabVIEW_Pompa 3"
   SymbolLibrary "Symbol library_18" at 361,151 size 16x15
      Appearance <- "OPC - do LabVIEW_Pompa 3"
   SymbolLibrary "Symbol library_19" at 408,166 size 28x45
      Appearance <- "OPC - do LabVIEW_Pompa 4"
   SymbolLibrary "Symbol library_20" at 409,151 size 16x16
      Appearance <- "OPC - do LabVIEW_Pompa 4"
   SymbolLibrary "Symbol library_21" at 571,166 size 28x45
      Appearance <- "OPC - do LabVIEW_Pompa 5"
   SymbolLibrary "Symbol library_22" at 572,152 size 16x15
      Appearance <- "OPC - do LabVIEW_Pompa 5"
   SymbolLibrary "Symbol library_23" at 618,165 size 28x45
      Appearance <- "OPC - do LabVIEW_Pompa 6"
   SymbolLibrary "Symbol library_24" at 619,151 size 16x15
      Appearance <- "OPC - do LabVIEW_Pompa 6"
   SymbolLibrary "Symbol library_25" at 417,372 size 28x45
      Appearance <- "OPC - do LabVIEW_Pompa 8"
   SymbolLibrary "Symbol library_26" at 419,416 size 16x18
      Appearance <- "OPC - do LabVIEW_Pompa 8"
   Bar "Bar_4" at 284,259 size 68x113; MinimumValue 0; MaximumValue 300
      ProcessValue <- "OPC - z LabVIEW_Poziom zbiornik 4"
   SymbolLibrary "Symbol library_27" at 370,352 size 117x20
      Appearance <- "OPC - do LabVIEW_Grzałka 4"
   IOField "I/O field_7" at 374,266 size 48x31; FormatPattern 999
      ProcessValue <- "HMI komunikacja_Czas utrz T w Z4 (timer)"
   IOField "I/O field_8" at 374,308 size 70x31; FormatPattern 999.9
      ProcessValue <- "OPC - z LabVIEW_Temp cieczy w zb4"
   TextField "Text field_8" at 433,280 size 33x18; Text 'sek.'
   TextField "Text field_9" at 441,316 size 25x23; Text '℃'
   SymbolLibrary "Symbol library_28" at 362,209 size 16x51
      Appearance <- "OPC - do LabVIEW_Pompa 3"
   SymbolLibrary "Symbol library_29" at 410,210 size 16x51
      Appearance <- "OPC - do LabVIEW_Pompa 4"
   IOField "I/O field_9" at 90,178 size 59x31; FormatPattern 99.9
      ProcessValue <- "OPC - z LabVIEW_Temp P1"
   TextField "Text field_10" at 125,209 size 25x23; Text '℃'
   IOField "I/O field_10" at 229,178 size 59x31; FormatPattern 99.9
      ProcessValue <- "OPC - z LabVIEW_Temp P2"
   TextField "Text field_11" at 269,205 size 25x23; Text '℃'
   IOField "I/O field_11" at 300,178 size 59x31; FormatPattern 99.9
      ProcessValue <- "OPC - z LabVIEW_Temp P3"
   TextField "Text field_12" at 338,206 size 25x23; Text '℃'
   IOField "I/O field_12" at 440,178 size 59x31; FormatPattern 99.9
      ProcessValue <- "OPC - z LabVIEW_Temp P4"
   TextField "Text field_13" at 476,205 size 25x23; Text '℃'
   IOField "I/O field_13" at 510,178 size 59x31; FormatPattern 99.9
      ProcessValue <- "OPC - z LabVIEW_Temp P5"
   TextField "Text field_14" at 547,206 size 25x23; Text '℃'
   IOField "I/O field_14" at 649,178 size 59x31; FormatPattern 99.9
      ProcessValue <- "OPC - z LabVIEW_Temp P6"
   TextField "Text field_15" at 684,206 size 25x23; Text '℃'
   IOField "I/O field_15" at 450,379 size 59x31; FormatPattern 99.9
      ProcessValue <- "OPC - z LabVIEW_Temp P8"
   TextField "Text field_16" at 508,391 size 25x23; Text '℃'
   IOField "I/O field_16" at 282,379 size 59x31; FormatPattern 99.9
      ProcessValue <- "OPC - z LabVIEW_Temp P7"
   TextField "Text field_17" at 338,388 size 25x23; Text '℃'
   TextField "Text field_18" at 217,156 size 78x21; Text 'Temp. P2'
   TextField "Text field_19" at 70,156 size 78x21; Text 'Temp. P1'
   TextField "Text field_20" at 428,156 size 78x21; Text 'Temp. P4'
   TextField "Text field_21" at 288,156 size 78x21; Text 'Temp. P3'
   TextField "Text field_22" at 501,156 size 78x21; Text 'Temp. P5'
   TextField "Text field_23" at 438,410 size 78x21; Text 'Temp. P8'
   TextField "Text field_24" at 638,155 size 78x21; Text 'Temp. P6'
   TextField "Text field_25" at 283,411 size 78x21; Text 'Temp. P7'
   TextField "Text field_26" at 104,39 size 23x97; Text 'Zbiornik 1'
   TextField "Text field_27" at 314,39 size 23x97; Text 'Zbiornik 2'
   TextField "Text field_28" at 524,39 size 23x97; Text 'Zbiornik 3'
   TextField "Text field_29" at 204,269 size 23x97; Text 'Zbiornik 4'
   SymbolLibrary "Symbol library_31" at 574,210 size 15x15
      Appearance <- "OPC - do LabVIEW_Pompa 5"
   Group "Group_1" at 588,210 size 48x29
   Group "Group" at 486,224 size 104x35
   Group "Group_3" at 199,224 size 104x35
   SymbolLibrary "Symbol library_34" at 200,210 size 15x15
      Appearance <- "OPC - do LabVIEW_Pompa 2"
   Group "Group_2" at 153,210 size 48x29
   SymbolLibrary "Symbol library_44" at 393,373 size 19x37
      Appearance <- "OPC - do LabVIEW_Zawór spustowy Z4"
   SymbolLibrary "Symbol library_45" at 599,151 size 19x37
      Appearance <- "OPC - do LabVIEW_Zawór spustowy Z3"
   SymbolLibrary "Symbol library_46" at 179,150 size 19x37
      Appearance <- "OPC - do LabVIEW_Zawór spustowy Z1"
   SymbolLibrary "Symbol library_47" at 389,150 size 19x37
      Appearance <- "OPC - do LabVIEW_Zawór spustowy Z2"
   Circle "Circle_1" at 33,298 size 48x48
      Appearance <- "HMI komunikacja_Blokada zmiany par. PRO"
   TextField "Text field_30" at 13,260 size 172x38; Text 'Możliwa zmiana parametrów procesu.'
   SymbolLibrary "Symbol library_30" at 606,210 size 30x29
      Appearance <- "OPC - do LabVIEW_Pompa 6"
   SymbolLibrary "Symbol library_32" at 588,224 size 31x15
      Appearance <- "OPC - do LabVIEW_Pompa 6"
   SymbolLibrary "Symbol library_33" at 566,224 size 24x15
      Appearance <- "HMI komunikacja_rura blue P5 i P6"
   SymbolLibrary "Symbol library_37" at 516,224 size 51x15
      Appearance <- "HMI komunikacja_rura blue P5 i P6"
   SymbolLibrary "Symbol library_39" at 486,224 size 31x29
      Appearance <- "HMI komunikacja_rura blue P5 i P6"
   SymbolLibrary "Symbol library_40" at 486,244 size 16x15
      Appearance <- "HMI komunikacja_rura blue P5 i P6"
   SymbolLibrary "Symbol library_35" at 153,210 size 30x29
      Appearance <- "OPC - do LabVIEW_Pompa 1"
   SymbolLibrary "Symbol library_36" at 170,224 size 31x15
      Appearance <- "OPC - do LabVIEW_Pompa 1"
   SymbolLibrary "Symbol library_38" at 199,224 size 24x15
      Appearance <- "HMI komunikacja_rura blue P1 i P2"
   SymbolLibrary "Symbol library_41" at 222,224 size 51x15
      Appearance <- "HMI komunikacja_rura blue P1 i P2"
   SymbolLibrary "Symbol library_42" at 272,224 size 31x29
      Appearance <- "HMI komunikacja_rura blue P1 i P2"
   SymbolLibrary "Symbol library_43" at 287,244 size 16x15
      Appearance <- "HMI komunikacja_rura blue P1 i P2"

